(* Logix 5000 project; controller Seperator 1756-L85E rev 33.11; software revision 33.01; part 6 of 7 *)
(* tags used below, declared in another part *)
   Bottle_Clamp_Pressure_actual_1 : REAL;
   Bottle_Clamp_Pressure_SP_1 : REAL;
   Bottle_level_actual_1 : REAL;
   Bottle_Slow_Fill_SP_1 : REAL;
   Bottle_Stop_Fill_SP_1 : REAL;
   Filling_Head_Sequencer_1 : DINT;
   Pump_Running_1 : BOOL;
   Aborted : SFC_STEP;
   bottle_clamp_out_delayF2 : TIMER;
   bottle_clamp_out_delayF3 : TIMER;
   Capper_Head_Sequencer : DINT;
   Comms_OK : BOOL;
   esd : BOOL;
   FC01 : FTV_ctrl;
   FI101 : REAL;
   FI101_Moving_Analog : Moving_Analog_Indicator;
   FI102 : REAL;
   FI102_Moving_Analog : Moving_Analog_Indicator;
   Filler_Index_complete : BOOL;
   Filling_Nozzle_Down_Delay2 : TIMER;
   Filling_Nozzle_Down_Delay3 : TIMER;
   Filling_Nozzle_up_Delay2 : TIMER;
   Filling_Nozzle_up_Delay3 : TIMER;
   Idle : SFC_STEP;
   II101 : REAL;
   II101_Moving_Analog : Moving_Analog_Indicator;
   Led_Code : INT;
   LI101 : REAL;
   LI101_Moving_Analog : Moving_Analog_Indicator;
   Main_Sequencer : DINT;
   Operator_Mode : BOOL;
   Phase_Control : Phase_Control;
   Phase_Result : DINT;
   PI102 : REAL;
   PI102_Moving_Analog : Moving_Analog_Indicator;
   Qtr_Sec_PLs : TIMER;
   Seperator_Control : PHASE;
   Seperator_State : BOOL[32];
   Status_Code : INT;
   Stopped : SFC_STEP;
   TI101 : REAL;
   TI101_Moving_Analog : Moving_Analog_Indicator;
   VI101 : REAL;
   VI101_Moving_Analog : Moving_Analog_Indicator;
(* Filler_Heads1, continued *)

ROUTINE Head_HMI_Collation   (* ladder *)
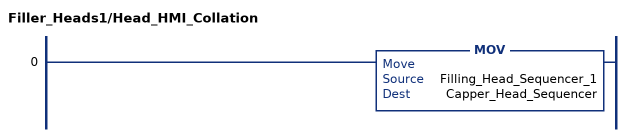
   0: MOV(Filling_Head_Sequencer_1,Capper_Head_Sequencer);
END_ROUTINE

ROUTINE Initialisation   (* ladder *)
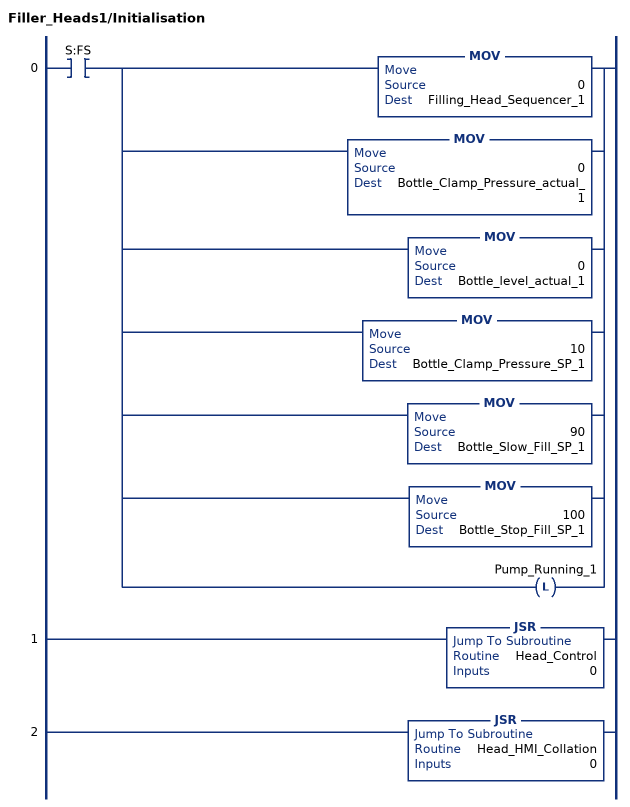
   0: XIC(S:FS)[MOV(0,Filling_Head_Sequencer_1) ,MOV(0,Bottle_Clamp_Pressure_actual_1) ,MOV(0,Bottle_level_actual_1) ,MOV(10,Bottle_Clamp_Pressure_SP_1) ,MOV(90,Bottle_Slow_Fill_SP_1) ,MOV(100,Bottle_Stop_Fill_SP_1) ,OTL(Pump_Running_1) ];
   1: JSR(Head_Control,0);
   2: JSR(Head_HMI_Collation,0);
END_ROUTINE
END_PROGRAM

PROGRAM Filler_Heads2   (* main routine Initialisation *)
VAR
   Alias_Head_Clamp_Pressure_SP_2 : ALIAS FOR Head_Clamp_Pressure_SP_2;
   Bottle_Clamp_Pressure_actual_2 : REAL := 10.799999;
   Bottle_Clamp_Pressure_SP_2 : REAL := 9.95;
   Bottle_Fill_Stop_SP_2 : REAL := 100.0;
   Bottle_level_actual_2 : REAL := 9.4;
   Bottle_Slow_Fill_SP_2 : REAL := 90.0;
   Filling_Head_Sequencer_2 : DINT := 3;
   Head1_98_Percent_temperatureSP_2 : REAL := 176.4;
   Head_Clamp_Pressure_SP_2 : REAL := 90.0;
   Head_Down_2 : BOOL;
   Head_Down_Stage1_2 : REAL := 18.0;
   Head_Down_Stage2_2 : REAL := 27.0;
   Head_Injection_Pressure_SP_2 : REAL := 75.0;
   Head_Injection_Stage1_2 : REAL := 18.75;
   Head_Injection_Stage2_2 : REAL := 33.75;
   Head_Injector_out_delay_2 : TIMER := (PRE := 2000);
   Head_moving_Down_2 : BOOL := 1;
   Head_moving_Up_2 : BOOL;
   Head_Up_2 : BOOL;
   Head_up_delay_2 : TIMER := (PRE := 2000);
   Pump_Running_2 : BOOL := 1;
   Rotary_Moulder_Head_Name_2 : STRING := 'Head 1'; {constant, access None}
   ScratchPad1_2 : REAL := 0.9;
   ScratchPad2_2 : REAL := 0.9;
   ScratchPad3_2 : REAL := 0.75;
   ScratchPad4_2 : REAL := 0.75;
   ScratchPad5_2 : REAL := 3.6;
   ScratchPad6_2 : REAL;
END_VAR

ROUTINE Head_Control   (* ladder *)
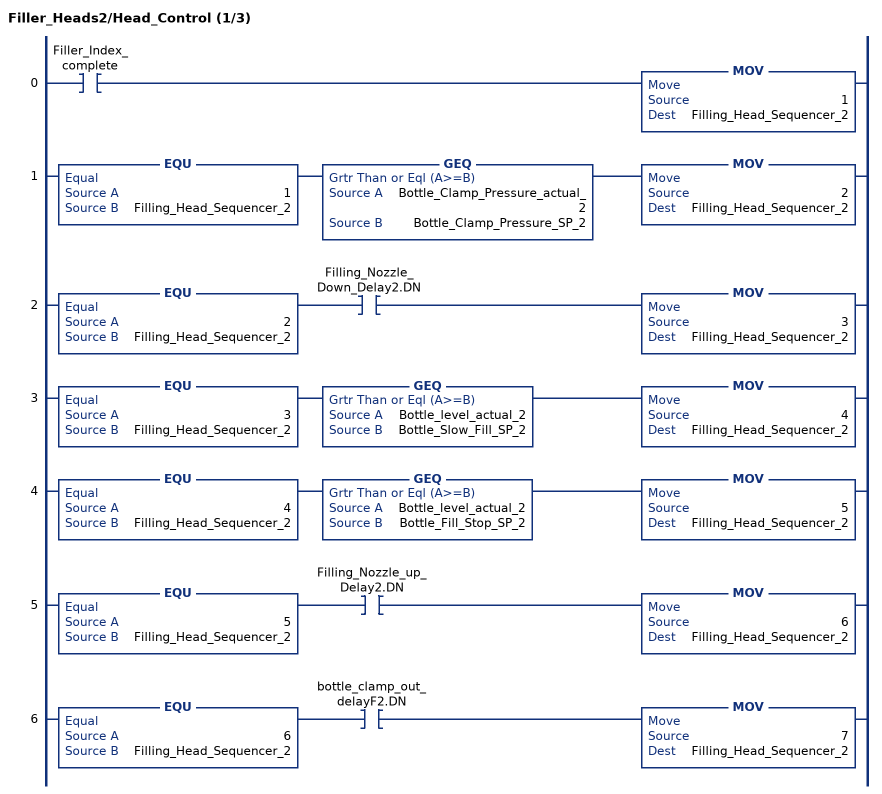
   0: XIC(Filler_Index_complete)MOV(1,Filling_Head_Sequencer_2);
   1: EQU(1,Filling_Head_Sequencer_2)GEQ(Bottle_Clamp_Pressure_actual_2,Bottle_Clamp_Pressure_SP_2)MOV(2,Filling_Head_Sequencer_2);
   2: EQU(2,Filling_Head_Sequencer_2)XIC(Filling_Nozzle_Down_Delay2.DN)MOV(3,Filling_Head_Sequencer_2);
   3: EQU(3,Filling_Head_Sequencer_2)GEQ(Bottle_level_actual_2,Bottle_Slow_Fill_SP_2)MOV(4,Filling_Head_Sequencer_2);
   4: EQU(4,Filling_Head_Sequencer_2)GEQ(Bottle_level_actual_2,Bottle_Fill_Stop_SP_2)MOV(5,Filling_Head_Sequencer_2);
   5: EQU(5,Filling_Head_Sequencer_2)XIC(Filling_Nozzle_up_Delay2.DN)MOV(6,Filling_Head_Sequencer_2);
   6: EQU(6,Filling_Head_Sequencer_2)XIC(bottle_clamp_out_delayF2.DN)MOV(7,Filling_Head_Sequencer_2);
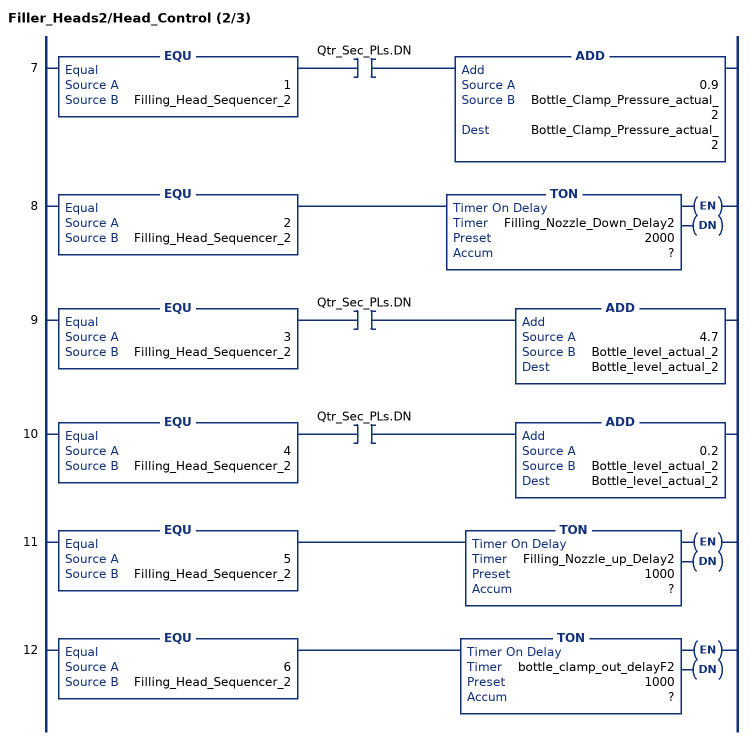
   7: EQU(1,Filling_Head_Sequencer_2)XIC(Qtr_Sec_PLs.DN)ADD(0.9,Bottle_Clamp_Pressure_actual_2,Bottle_Clamp_Pressure_actual_2);
   8: EQU(2,Filling_Head_Sequencer_2)TON(Filling_Nozzle_Down_Delay2,?,?);
   9: EQU(3,Filling_Head_Sequencer_2)XIC(Qtr_Sec_PLs.DN)ADD(4.7,Bottle_level_actual_2,Bottle_level_actual_2);
   10: EQU(4,Filling_Head_Sequencer_2)XIC(Qtr_Sec_PLs.DN)ADD(0.2,Bottle_level_actual_2,Bottle_level_actual_2);
   11: EQU(5,Filling_Head_Sequencer_2)TON(Filling_Nozzle_up_Delay2,?,?);
   12: EQU(6,Filling_Head_Sequencer_2)TON(bottle_clamp_out_delayF2,?,?);
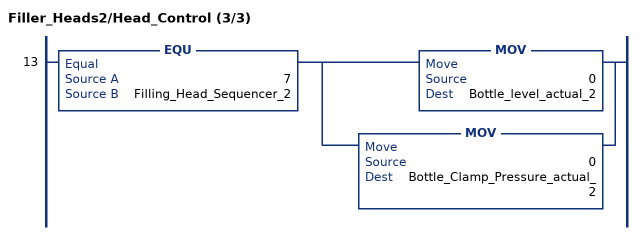
   13: EQU(7,Filling_Head_Sequencer_2)[MOV(0,Bottle_level_actual_2) ,MOV(0,Bottle_Clamp_Pressure_actual_2) ];
END_ROUTINE

ROUTINE Head_HMI_Collation   (* ladder *)
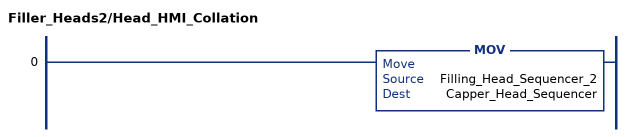
   0: MOV(Filling_Head_Sequencer_2,Capper_Head_Sequencer);
END_ROUTINE

ROUTINE Initialisation   (* ladder *)
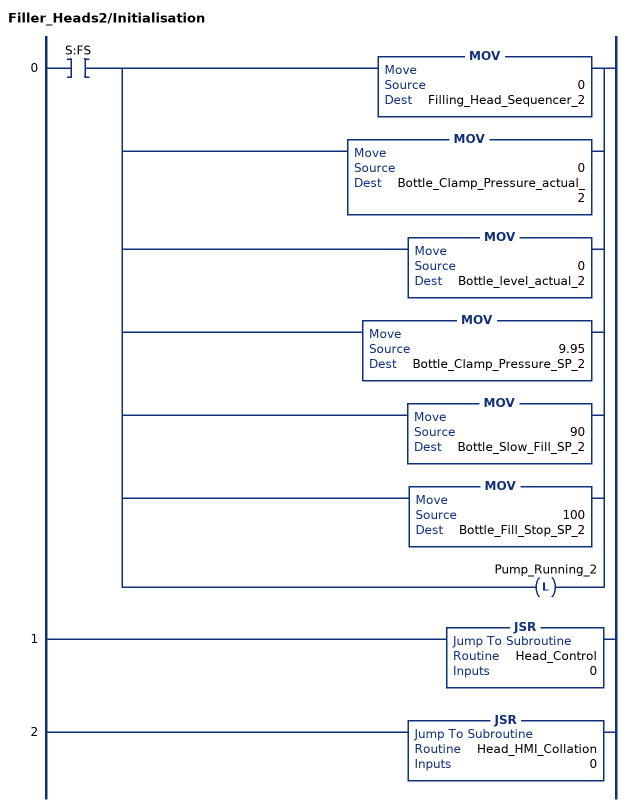
   0: XIC(S:FS)[MOV(0,Filling_Head_Sequencer_2) ,MOV(0,Bottle_Clamp_Pressure_actual_2) ,MOV(0,Bottle_level_actual_2) ,MOV(9.95,Bottle_Clamp_Pressure_SP_2) ,MOV(90,Bottle_Slow_Fill_SP_2) ,MOV(100,Bottle_Fill_Stop_SP_2) ,OTL(Pump_Running_2) ];
   1: JSR(Head_Control,0);
   2: JSR(Head_HMI_Collation,0);
END_ROUTINE
END_PROGRAM

PROGRAM Filler_Heads3   (* main routine Initialisation *)
VAR
   Alias_Head_Clamp_Pressure_SP_3 : ALIAS FOR Head_Clamp_Pressure_SP_3;
   Bottle_Clamp_Pressure_actual_3 : REAL := 10.799999;
   Bottle_Clamp_Pressure_SP_3 : REAL := 9.97;
   Bottle_Fill_Stop_SP_3 : REAL := 100.0;
   Bottle_level_actual_3 : REAL := 14.099999;
   Bottle_Slow_Fill_SP_3 : REAL := 90.0;
   Filling_Head_Sequencer_3 : DINT := 3;
   Head1_98_Percent_temperatureSP_3 : REAL := 176.4;
   Head_Clamp_Pressure_SP_3 : REAL := 90.0;
   Head_Down_3 : BOOL;
   Head_Down_Stage1_3 : REAL := 18.0;
   Head_Down_Stage2_3 : REAL := 27.0;
   Head_Injection_Pressure_SP_3 : REAL := 75.0;
   Head_Injection_Stage1_3 : REAL := 18.75;
   Head_Injection_Stage2_3 : REAL := 33.75;
   Head_Injector_out_delay_3 : TIMER := (PRE := 2000);
   Head_moving_Down_3 : BOOL := 1;
   Head_moving_Up_3 : BOOL;
   Head_Up_3 : BOOL;
   Head_up_delay_3 : TIMER := (PRE := 2000);
   Pump_Running_3 : BOOL := 1;
   Rotary_Moulder_Head_Name_3 : STRING := 'Head 1'; {constant, access None}
   ScratchPad1_3 : REAL := 0.9;
   ScratchPad2_3 : REAL := 0.9;
   ScratchPad3_3 : REAL := 0.75;
   ScratchPad4_3 : REAL := 0.75;
   ScratchPad5_3 : REAL := 3.6;
   ScratchPad6_3 : REAL;
END_VAR

ROUTINE Head_Control   (* ladder *)
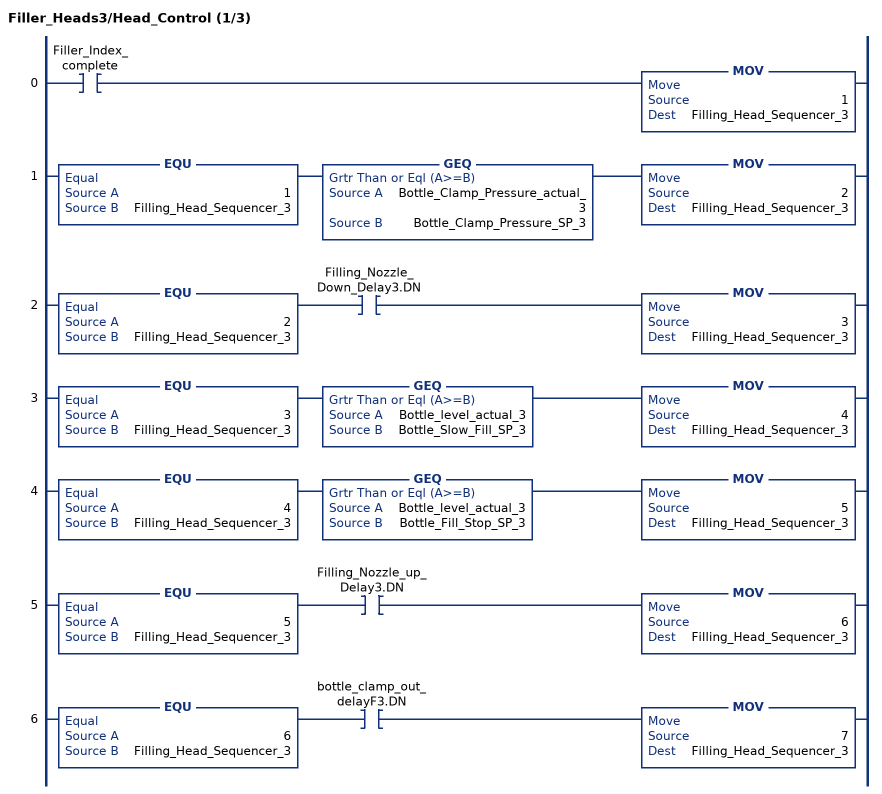
   0: XIC(Filler_Index_complete)MOV(1,Filling_Head_Sequencer_3);
   1: EQU(1,Filling_Head_Sequencer_3)GEQ(Bottle_Clamp_Pressure_actual_3,Bottle_Clamp_Pressure_SP_3)MOV(2,Filling_Head_Sequencer_3);
   2: EQU(2,Filling_Head_Sequencer_3)XIC(Filling_Nozzle_Down_Delay3.DN)MOV(3,Filling_Head_Sequencer_3);
   3: EQU(3,Filling_Head_Sequencer_3)GEQ(Bottle_level_actual_3,Bottle_Slow_Fill_SP_3)MOV(4,Filling_Head_Sequencer_3);
   4: EQU(4,Filling_Head_Sequencer_3)GEQ(Bottle_level_actual_3,Bottle_Fill_Stop_SP_3)MOV(5,Filling_Head_Sequencer_3);
   5: EQU(5,Filling_Head_Sequencer_3)XIC(Filling_Nozzle_up_Delay3.DN)MOV(6,Filling_Head_Sequencer_3);
   6: EQU(6,Filling_Head_Sequencer_3)XIC(bottle_clamp_out_delayF3.DN)MOV(7,Filling_Head_Sequencer_3);
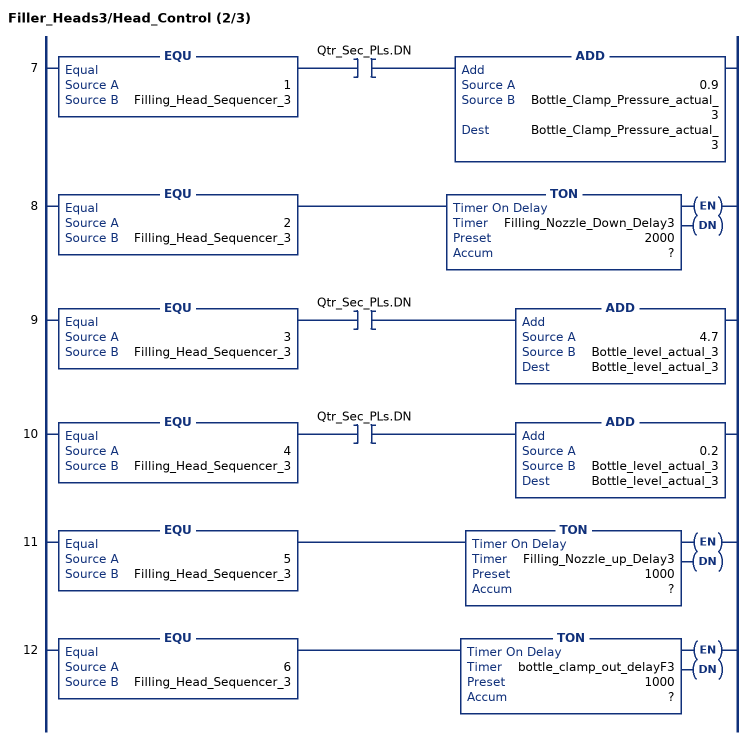
   7: EQU(1,Filling_Head_Sequencer_3)XIC(Qtr_Sec_PLs.DN)ADD(0.9,Bottle_Clamp_Pressure_actual_3,Bottle_Clamp_Pressure_actual_3);
   8: EQU(2,Filling_Head_Sequencer_3)TON(Filling_Nozzle_Down_Delay3,?,?);
   9: EQU(3,Filling_Head_Sequencer_3)XIC(Qtr_Sec_PLs.DN)ADD(4.7,Bottle_level_actual_3,Bottle_level_actual_3);
   10: EQU(4,Filling_Head_Sequencer_3)XIC(Qtr_Sec_PLs.DN)ADD(0.2,Bottle_level_actual_3,Bottle_level_actual_3);
   11: EQU(5,Filling_Head_Sequencer_3)TON(Filling_Nozzle_up_Delay3,?,?);
   12: EQU(6,Filling_Head_Sequencer_3)TON(bottle_clamp_out_delayF3,?,?);
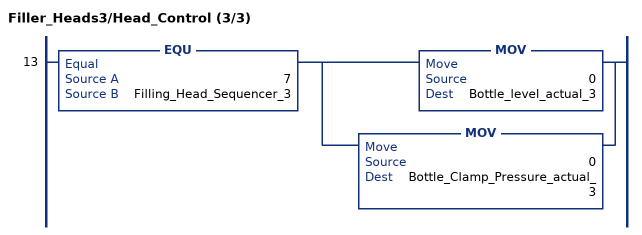
   13: EQU(7,Filling_Head_Sequencer_3)[MOV(0,Bottle_level_actual_3) ,MOV(0,Bottle_Clamp_Pressure_actual_3) ];
END_ROUTINE

ROUTINE Head_HMI_Collation   (* ladder *)
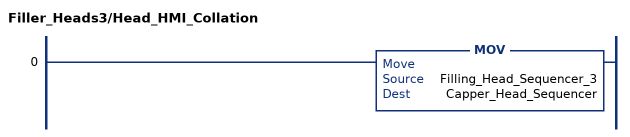
   0: MOV(Filling_Head_Sequencer_3,Capper_Head_Sequencer);
END_ROUTINE

ROUTINE Initialisation   (* ladder *)
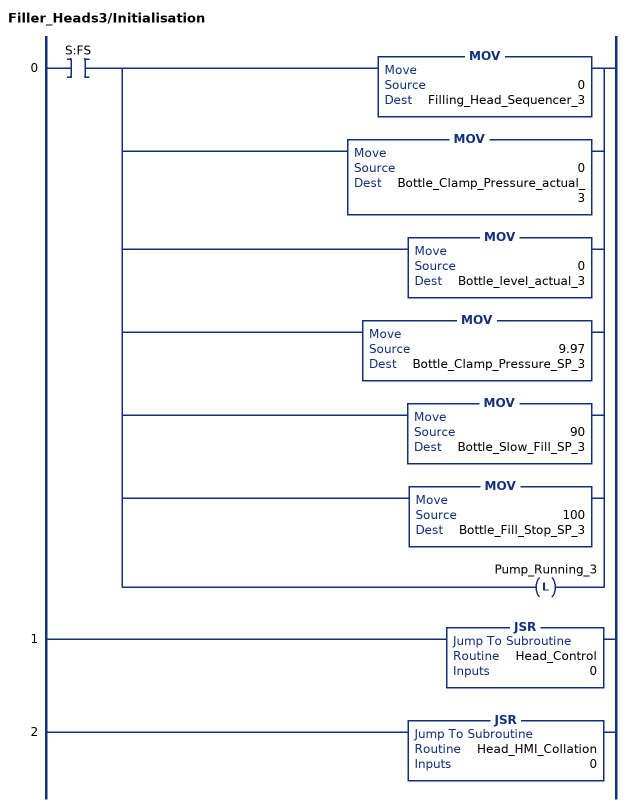
   0: XIC(S:FS)[MOV(0,Filling_Head_Sequencer_3) ,MOV(0,Bottle_Clamp_Pressure_actual_3) ,MOV(0,Bottle_level_actual_3) ,MOV(9.97,Bottle_Clamp_Pressure_SP_3) ,MOV(90,Bottle_Slow_Fill_SP_3) ,MOV(100,Bottle_Fill_Stop_SP_3) ,OTL(Pump_Running_3) ];
   1: JSR(Head_Control,0);
   2: JSR(Head_HMI_Collation,0);
END_ROUTINE
END_PROGRAM

PROGRAM IO_Simulation   (* main routine MainRoutine *)
VAR
   djw : BOOL;
   DwellTimer : TIMER[32];
   RunSEQ : DINT[4];
   StopSEQ : DINT[4];
END_VAR

ROUTINE Leds_Control   (* ladder *)
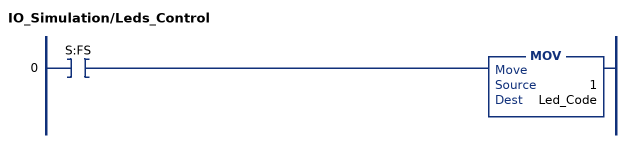
   0: XIC(S:FS)MOV(1,Led_Code);
END_ROUTINE

ROUTINE MainRoutine   (* ladder *)
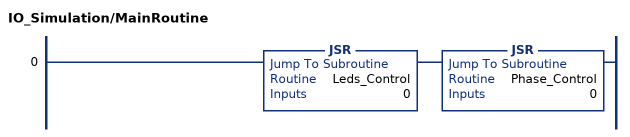
   0: JSR(Leds_Control,0)JSR(Phase_Control,0);
END_ROUTINE

ROUTINE Phase_Control   (* ladder *)
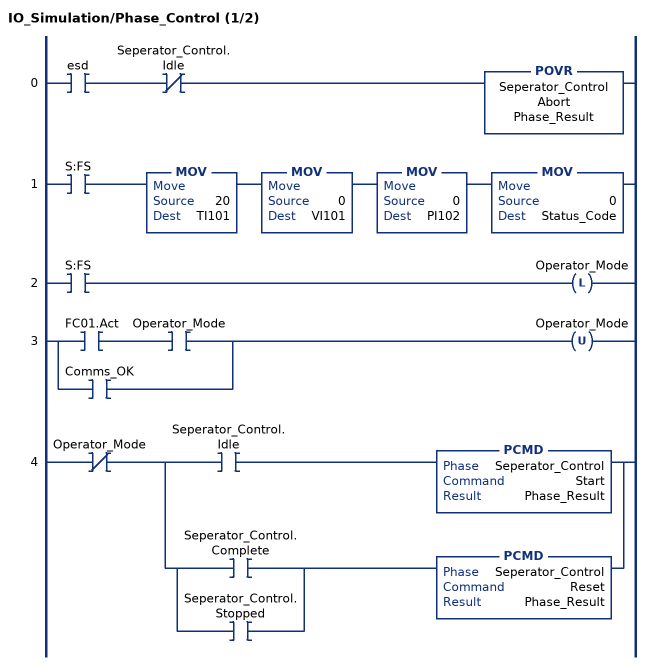
   0: XIC(esd)XIO(Seperator_Control.Idle)POVR(Seperator_Control,Abort,Phase_Result);
   1: XIC(S:FS)MOV(20,TI101)MOV(0,VI101)MOV(0,PI102)MOV(0,Status_Code);
   2: XIC(S:FS)OTL(Operator_Mode);
   3: [XIC(FC01.Act) XIC(Operator_Mode) ,XIC(Comms_OK) ]OTU(Operator_Mode);
   4: XIO(Operator_Mode)[XIC(Seperator_Control.Idle) PCMD(Seperator_Control,Start,Phase_Result) ,[XIC(Seperator_Control.Complete) ,XIC(Seperator_Control.Stopped) ] PCMD(Seperator_Control,Reset,Phase_Result) ];
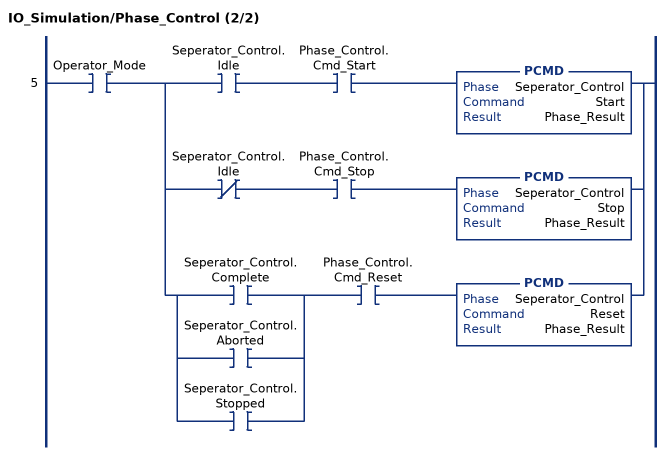
   5: XIC(Operator_Mode)[XIC(Seperator_Control.Idle) XIC(Phase_Control.Cmd_Start) PCMD(Seperator_Control,Start,Phase_Result) ,XIO(Seperator_Control.Idle) XIC(Phase_Control.Cmd_Stop) PCMD(Seperator_Control,Stop,Phase_Result) ,[[XIC(Seperator_Control.Complete) ,XIC(Seperator_Control.Aborted) ] ,XIC(Seperator_Control.Stopped) ] XIC(Phase_Control.Cmd_Reset) PCMD(Seperator_Control,Reset,Phase_Result) ];
END_ROUTINE
END_PROGRAM

PROGRAM Main_Sequencer   (* main routine Main_Sequencer *)
VAR
   Empty_Vacuum_Silo1_ons : BOOL := 1;
   Empty_Vacuum_Silo2_ons : BOOL;
   Empty_Vacuum_Silo3_ons : BOOL := 1;
   Empty_Vacuum_Silo4_ons : BOOL;
   Fill_Vacuum_Silo1_ons : BOOL := 1;
   Fill_Vacuum_Silo2_ons : BOOL;
   Fill_Vacuum_Silo3_ons : BOOL;
   Fill_Vacuum_Silo4_ons : BOOL;
   Fill_Vacuum_Silo_ons : BOOL;
   Run_Vacuum_Silo_Decision_Manager : BOOL := 1;
END_VAR

ROUTINE HMI_collation   (* ladder *)
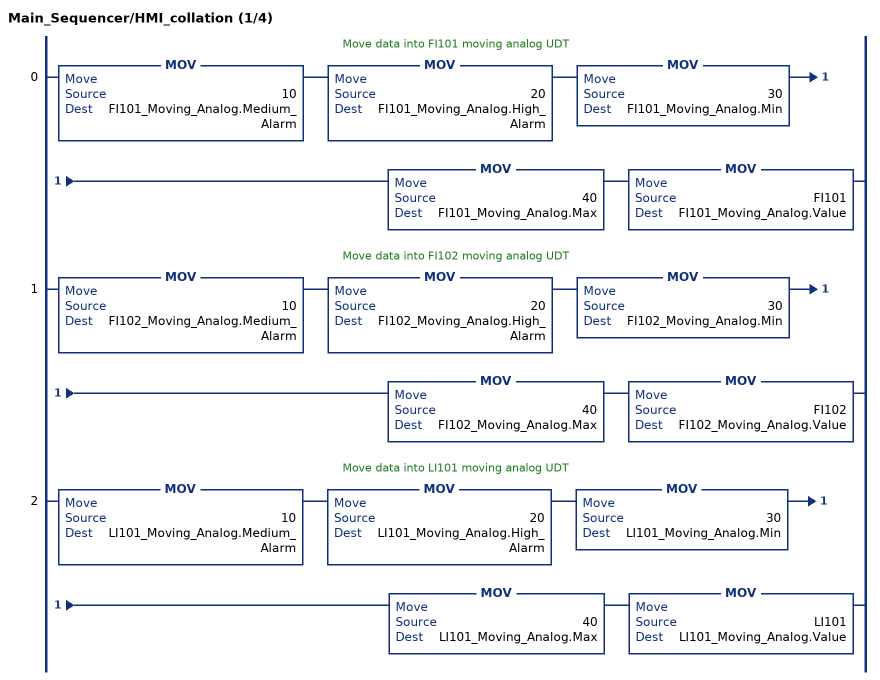
   // Move data into FI101 moving analog UDT
   0: MOV(10,FI101_Moving_Analog.Medium_Alarm)MOV(20,FI101_Moving_Analog.High_Alarm)MOV(30,FI101_Moving_Analog.Min)MOV(40,FI101_Moving_Analog.Max)MOV(FI101,FI101_Moving_Analog.Value);
   // Move data into FI102 moving analog UDT
   1: MOV(10,FI102_Moving_Analog.Medium_Alarm)MOV(20,FI102_Moving_Analog.High_Alarm)MOV(30,FI102_Moving_Analog.Min)MOV(40,FI102_Moving_Analog.Max)MOV(FI102,FI102_Moving_Analog.Value);
   // Move data into LI101 moving analog UDT
   2: MOV(10,LI101_Moving_Analog.Medium_Alarm)MOV(20,LI101_Moving_Analog.High_Alarm)MOV(30,LI101_Moving_Analog.Min)MOV(40,LI101_Moving_Analog.Max)MOV(LI101,LI101_Moving_Analog.Value);
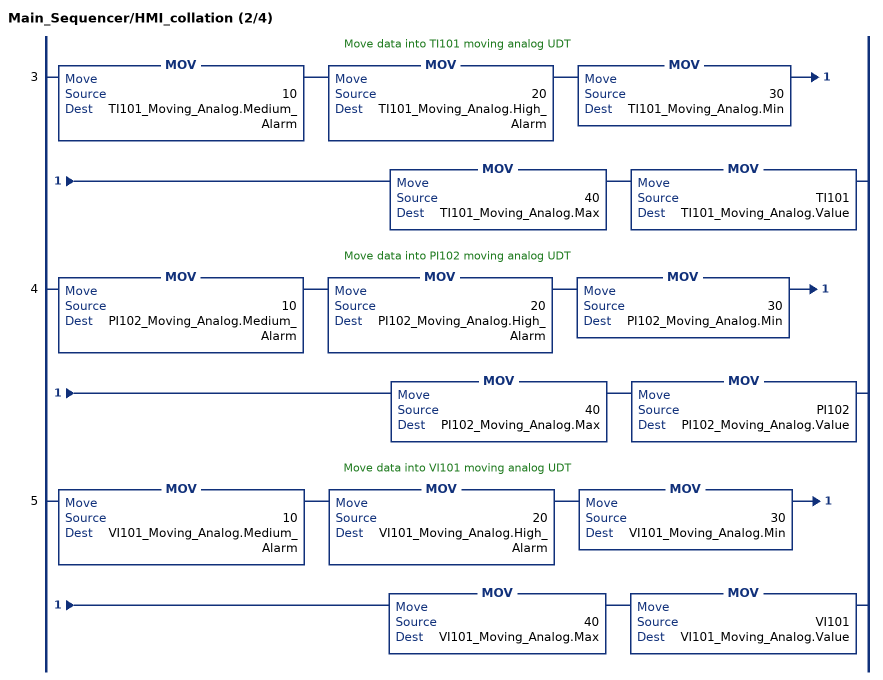
   // Move data into TI101 moving analog UDT
   3: MOV(10,TI101_Moving_Analog.Medium_Alarm)MOV(20,TI101_Moving_Analog.High_Alarm)MOV(30,TI101_Moving_Analog.Min)MOV(40,TI101_Moving_Analog.Max)MOV(TI101,TI101_Moving_Analog.Value);
   // Move data into PI102 moving analog UDT
   4: MOV(10,PI102_Moving_Analog.Medium_Alarm)MOV(20,PI102_Moving_Analog.High_Alarm)MOV(30,PI102_Moving_Analog.Min)MOV(40,PI102_Moving_Analog.Max)MOV(PI102,PI102_Moving_Analog.Value);
   // Move data into VI101 moving analog UDT
   5: MOV(10,VI101_Moving_Analog.Medium_Alarm)MOV(20,VI101_Moving_Analog.High_Alarm)MOV(30,VI101_Moving_Analog.Min)MOV(40,VI101_Moving_Analog.Max)MOV(VI101,VI101_Moving_Analog.Value);
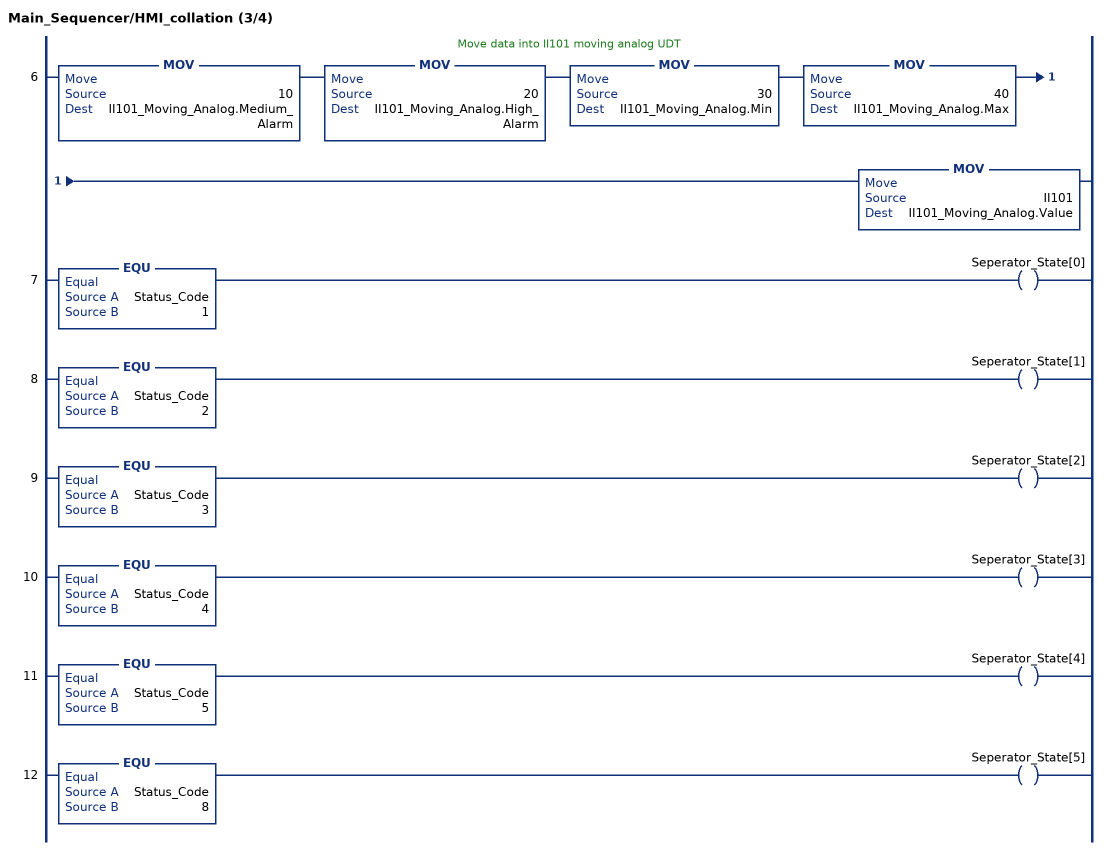
   // Move data into II101 moving analog UDT
   6: MOV(10,II101_Moving_Analog.Medium_Alarm)MOV(20,II101_Moving_Analog.High_Alarm)MOV(30,II101_Moving_Analog.Min)MOV(40,II101_Moving_Analog.Max)MOV(II101,II101_Moving_Analog.Value);
   7: EQU(Status_Code,1)OTE(Seperator_State[0]);
   8: EQU(Status_Code,2)OTE(Seperator_State[1]);
   9: EQU(Status_Code,3)OTE(Seperator_State[2]);
   10: EQU(Status_Code,4)OTE(Seperator_State[3]);
   11: EQU(Status_Code,5)OTE(Seperator_State[4]);
   12: EQU(Status_Code,8)OTE(Seperator_State[5]);
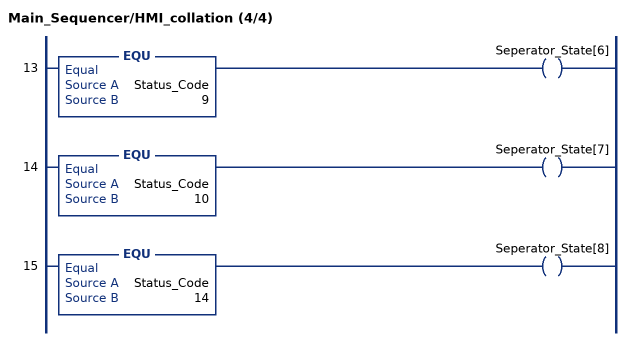
   13: EQU(Status_Code,9)OTE(Seperator_State[6]);
   14: EQU(Status_Code,10)OTE(Seperator_State[7]);
   15: EQU(Status_Code,14)OTE(Seperator_State[8]);
END_ROUTINE
